// TIA Portal project "TestEssProtoFreia" (V13) (continued)

         AN    "ASCOenManuel";
         =     "PLC_to_Epics".CV550.sAuto;
END_REGION

REGION Network 13: spare - VB chan 7
   RUNG wire#powerrail
      Contact( "voie 7 chaufferette BV" )
      Coil( "PLC_to_Epics"."spare-VB-7".sHtrOn )
   END_RUNG
   // the same network as SCL:
   "PLC_to_Epics"."spare-VB-7".sHtrOn := "voie 7 chaufferette BV";
END_REGION

REGION Network 14: spare - VB chan 8
   RUNG wire#powerrail
      Contact( "voie 8 chaufferette BV" )
      Coil( "PLC_to_Epics"."spare-VB-8".sHtrOn )
   END_RUNG
   // the same network as SCL:
   "PLC_to_Epics"."spare-VB-8".sHtrOn := "voie 8 chaufferette BV";
END_REGION

REGION Network 15: spare VB chan 9
   RUNG wire#powerrail
      Contact( "voie 9 chaufferette BV" )
      Coil( "PLC_to_Epics"."spare-VB-9".sHtrOn )
   END_RUNG
   // the same network as SCL:
   "PLC_to_Epics"."spare-VB-9".sHtrOn := "voie 9 chaufferette BV";
END_REGION

REGION Network 16: spare - VB chan 10
   RUNG wire#powerrail
      Contact( "voie 10  chaufferette BV" )
      Coil( "PLC_to_Epics"."spare-VB-10".sHtrOn )
   END_RUNG
   // the same network as SCL:
   "PLC_to_Epics"."spare-VB-10".sHtrOn := "voie 10  chaufferette BV";
END_REGION

REGION Network 17: spare - VB chan 11
   RUNG wire#powerrail
      Contact( "voie 11 chaufferette BV" )
      Coil( "PLC_to_Epics"."spare-VB-11".sHtrOn )
   END_RUNG
   // the same network as SCL:
   "PLC_to_Epics"."spare-VB-11".sHtrOn := "voie 11 chaufferette BV";
END_REGION

REGION Network 18: EH901-902 CM chan 1
   RUNG wire#powerrail
      Contact( "voie 1 chaufferette CM" )
      Coil( "PLC_to_Epics"."EH901-902".sHtrOn )
   END_RUNG
   // the same network as SCL:
   "PLC_to_Epics"."EH901-902".sHtrOn := "voie 1 chaufferette CM";
END_REGION

REGION Network 19: EH913-914 CM channel 4
   RUNG wire#powerrail
      Contact( "voie 4 chaufferette CM" )
      Coil( "PLC_to_Epics"."EH913-914".sHtrOn )
   END_RUNG
   // the same network as SCL:
   "PLC_to_Epics"."EH913-914".sHtrOn := "voie 4 chaufferette CM";
END_REGION

REGION Network 20: EH933-934 - CM chan 5
   RUNG wire#powerrail
      Contact( "voie 5 chaufferette CM" )
      Coil( "PLC_to_Epics"."EH933-934".sHtrOn )
   END_RUNG
   // the same network as SCL:
   "PLC_to_Epics"."EH933-934".sHtrOn := "voie 5 chaufferette CM";
END_REGION

REGION Network 21: EH921 - CM chan 6
   RUNG wire#powerrail
      Contact( "voie 6 chaufferette CM" )
      Coil( "PLC_to_Epics".EH921.sHtrOn )
   END_RUNG
   // the same network as SCL:
   "PLC_to_Epics".EH921.sHtrOn := "voie 6 chaufferette CM";
END_REGION

REGION Network 22: EH931-932 - CM chan 7
   RUNG wire#powerrail
      Contact( "voie 7 chaufferette CM" )
      Coil( "PLC_to_Epics"."EH931-932".sHtrOn )
   END_RUNG
   // the same network as SCL:
   "PLC_to_Epics"."EH931-932".sHtrOn := "voie 7 chaufferette CM";
END_REGION

REGION Network 23: EH915-916 - CM chan 8
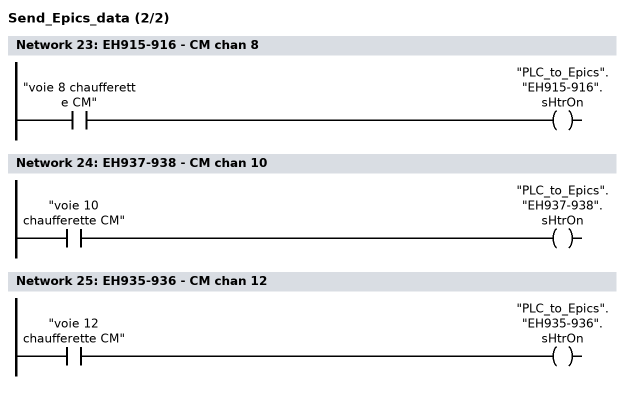
   RUNG wire#powerrail
      Contact( "voie 8 chaufferette CM" )
      Coil( "PLC_to_Epics"."EH915-916".sHtrOn )
   END_RUNG
   // the same network as SCL:
   "PLC_to_Epics"."EH915-916".sHtrOn := "voie 8 chaufferette CM";
END_REGION

REGION Network 24: EH937-938 - CM chan 10
   RUNG wire#powerrail
      Contact( "voie 10 chaufferette CM" )
      Coil( "PLC_to_Epics"."EH937-938".sHtrOn )
   END_RUNG
   // the same network as SCL:
   "PLC_to_Epics"."EH937-938".sHtrOn := "voie 10 chaufferette CM";
END_REGION

REGION Network 25: EH935-936 - CM chan 12
   RUNG wire#powerrail
      Contact( "voie 12 chaufferette CM" )
      Coil( "PLC_to_Epics"."EH935-936".sHtrOn )
   END_RUNG
   // the same network as SCL:
   "PLC_to_Epics"."EH935-936".sHtrOn := "voie 12 chaufferette CM";
END_REGION

REGION Network 26 (STL): Status bits
         A     "Graph/manuelle";
         =     "PLC_to_Epics".sManual;
         A     "ErreurSupervision";
         =     "PLC_to_Epics".sGrafcetERR;
         A     "Etat initial";
         =     "PLC_to_Epics".sGS1;
         A     "EtatCdtCryo";
         =     "PLC_to_Epics".sGS2;
         A     "EtatAttMef";
         =     "PLC_to_Epics".sGS3;
         A     "EtatMEFazote";
         =     "PLC_to_Epics".sGS4;
         A     "EtatMEFhelium";
         =     "PLC_to_Epics".sGS5;
         A     "EtatMode4k";
         =     "PLC_to_Epics".sGS6;
         A     "EtatModeStandBy";
         =     "PLC_to_Epics".sGS7;
         A     "EtatMode2K";
         =     "PLC_to_Epics".sGS8;
         A     "Etatrechauffage";
         =     "PLC_to_Epics".sGS10;
         A     "conditionTempMEFheliumOK";
         =     "PLC_to_Epics".sTransTempOK;
         A     "TransMode4K";
         =     "PLC_to_Epics".sTransMode4K;
         A     "EPICS_COMM_OK";
         =     "PLC_to_Epics".EpicsCommOK;
         A     "HNOSS_COMM_OK";
         =     "PLC_to_Epics".HNOSSCommOK;
END_REGION

REGION Network 27 (STL): Real parameters read-back (LHe level PID settings)
         L     "TriggerPIDcv01";
         T     "PLC_to_Epics".TrigPID_CV01.sSetV;
         L     "TriggerPIDcv02";
         T     "PLC_to_Epics".TrigPID_CV02.sSetV;
         L     "TriggerPIDcv03";
         T     "PLC_to_Epics".TrigPID_CV03.sSetV;
         L     "LT01LevelSP2k";
         T     "PLC_to_Epics".PID_LT01_CV01_SP.sSetV;
         L     "LT01LevelSP";
         T     "PLC_to_Epics".PID_LT01_CV02_SP.sSetV;
         L     "LT03LevelSP";
         T     "PLC_to_Epics".PID_LT03_CV03_SP.sSetV;
END_REGION

REGION Network 28 (STL): Real parameters read-back (CV550l PID settings)
         L     "RéguleASCO02_SP";
         T     "PLC_to_Epics".PID_PT01_CV550_SP.sSetV;
END_REGION
END_FUNCTION

FUNCTION "Cmds_from_Epics" : Void   // FC33, STL
TITLE = Process data from Epics
{ S7_Optimized_Access := 'FALSE' }
VERSION : 0.1
BEGIN

REGION Network 1: Switch to remote mode (control from Epics)
         A     "Epics_to_PLC".cmdRemoteMode;
         R     "LocalMode";
         R     "Epics_to_PLC".cmdRemoteMode;
END_REGION

REGION Network 2: If Local mode - return
         A     "LocalMode";
         SAVE;
         BEC;
END_REGION

REGION Network 3: Switch to local mode (control from Epics)
         A     "Epics_to_PLC".cmdLocalMode;
         S     "LocalMode";
         R     "Epics_to_PLC".cmdLocalMode;
END_REGION

REGION Network 4: If Local mode - return
         A     "LocalMode";
         SAVE;
         BEC;
END_REGION

REGION Network 5: Test data (copy block of data)
   //      OPN   "Epics_to_PLC"
   //      OPNDI "PLC_to_Epics"
   //      LAR1  P#12.0
   //      LAR2  P#12.0
   //      L     14
   //lp1:  T     #cnt
   //      L DBD [ AR1 , P#0.0 ]
   //      T DID [ AR2 , P#0.0 ]
   //      +AR1  P#4.0
   //      +AR2  P#4.0
   //      L     #cnt
   //      LOOP  lp1
END_REGION

REGION Network 6: CV01 Man/Auto
         A     "Epics_to_PLC".CV01.cmdAuto;
         R     "CV01_ManAuto";
         A     "Epics_to_PLC".CV01.cmdMan;
         S     "CV01_ManAuto";
END_REGION

REGION Network 7: CV01 - set Value
         A     "CV01_ManAuto";
         A     "Epics_to_PLC".CV01.cmdSet;
         JNB   Label_0;
         L     "Epics_to_PLC".CV01.cSetv;
         T     "CV01_HMI_VAL";
         SET;
         SAVE;
         CLR;
   Label_0:A     BR;
         R     "Epics_to_PLC".CV01.cmdSet;
END_REGION

REGION Network 8: CV02 Man/Auto
         A     "Epics_to_PLC".CV02.cmdAuto;
         R     "CV02_ManAuto";
         A     "Epics_to_PLC".CV02.cmdMan;
         S     "CV02_ManAuto";
END_REGION

REGION Network 9: CV02 - set Value
         A     "CV02_ManAuto";
         A     "Epics_to_PLC".CV02.cmdSet;
         JNB   Label_1;
         L     "Epics_to_PLC".CV02.cSetv;
         T     "CV02_HMI_VAL";
         SET;
         SAVE;
         CLR;
   Label_1:A     BR;
         R     "Epics_to_PLC".CV02.cmdSet;
END_REGION

REGION Network 10: CV03 Man/Auto
         A     "Epics_to_PLC".CV03.cmdAuto;
         R     "CV03_ManAuto";
         A     "Epics_to_PLC".CV03.cmdMan;
         S     "CV03_ManAuto";
END_REGION

REGION Network 11: CV03 - set Value
         A     "CV03_ManAuto";
         A     "Epics_to_PLC".CV03.cmdSet;
         JNB   Label_2;
         L     "Epics_to_PLC".CV03.cSetv;
         T     "CV03_HMI_VAL";
         SET;
         SAVE;
         CLR;
   Label_2:A     BR;
         R     "Epics_to_PLC".CV03.cmdSet;
END_REGION

REGION Network 12: CV04 Man/Auto
         A     "Epics_to_PLC".CV04.cmdAuto;
         R     "CV04_ManAuto";
         A     "Epics_to_PLC".CV04.cmdMan;
         S     "CV04_ManAuto";
END_REGION

REGION Network 13: CV04 - set Value
         A     "CV04_ManAuto";
         A     "Epics_to_PLC".CV04.cmdSet;
         JNB   Label_3;
         L     "Epics_to_PLC".CV04.cSetv;
         T     "CV04_HMI_VAL";
         SET;
         SAVE;
         CLR;
   Label_3:A     BR;
         R     "Epics_to_PLC".CV04.cmdSet;
END_REGION

REGION Network 14: CV05 Man/Auto
END_REGION

REGION Network 15: CV05 - set Value NOTE: NO LOCAL FALG !!!!!!!!!!!!!!!!!!!
         A     "Epics_to_PLC".CV05.cmdSet;
         JNB   Label_4;
         L     "Epics_to_PLC".CV05.cSetv;
         T     "CV05_HMI_VAL";
         SET;
         SAVE;
         CLR;
   Label_4:A     BR;
         R     "Epics_to_PLC".CV05.cmdSet;
END_REGION

REGION Network 16: CV07 Man/Auto
         A     "Epics_to_PLC".CV07.cmdAuto;
         R     "CV07_ManAuto";
         A     "Epics_to_PLC".CV07.cmdMan;
         S     "CV07_ManAuto";
END_REGION

REGION Network 17: CV07 - set Value
         A     "CV07_ManAuto";
         A     "Epics_to_PLC".CV07.cmdSet;
         JNB   Label_5;
         L     "Epics_to_PLC".CV07.cSetv;
         T     "CV07_HMI_VAL";
         SET;
         SAVE;
         CLR;
   Label_5:A     BR;
         R     "Epics_to_PLC".CV07.cmdSet;
END_REGION

REGION Network 18: CV60 Man/Auto
         A     "Epics_to_PLC".CV60.cmdAuto;
         R     "CV60_ManAuto";
         A     "Epics_to_PLC".CV60.cmdMan;
         S     "CV60_ManAuto";
END_REGION

REGION Network 19: CV60 - set Value
         A     "CV60_ManAuto";
         A     "Epics_to_PLC".CV60.cmdSet;
         JNB   Label_6;
         L     "Epics_to_PLC".CV60.cSetv;
         T     "CV60_HMI_VAL";
         SET;
         SAVE;
         CLR;
   Label_6:A     BR;
         R     "Epics_to_PLC".CV60.cmdSet;
END_REGION

REGION Network 20: CV61 Man/Auto
         A     "Epics_to_PLC".CV61.cmdAuto;
         R     "CV61_ManAuto";
         A     "Epics_to_PLC".CV61.cmdMan;
         S     "CV61_ManAuto";
END_REGION

REGION Network 21: CV61 - set Value
         A     "CV61_ManAuto";
         A     "Epics_to_PLC".CV61.cmdSet;
         JNB   Label_7;
         L     "Epics_to_PLC".CV61.cSetv;
         T     "CV61_HMI_VAL";
         SET;
         SAVE;
         CLR;
   Label_7:A     BR;
         R     "Epics_to_PLC".CV61.cmdSet;
END_REGION

REGION Network 22: CV62 Man/Auto
END_REGION

REGION Network 23: CV62 - set Value
         A     "Epics_to_PLC".CV62.cmdSet;
         JNB   Label_8;
         L     "Epics_to_PLC".CV62.cSetv;
         T     "CV62_HMI_VAL";
         SET;
         SAVE;
         CLR;
   Label_8:A     BR;
         R     "Epics_to_PLC".CV62.cmdSet;
END_REGION

REGION Network 24: CV550 Man/Auto
         A     "Epics_to_PLC".CV550.cmdAuto;
         R     "ASCOenManuel";
         A     "Epics_to_PLC".CV550.cmdMan;
         S     "ASCOenManuel";
END_REGION

REGION Network 25: CV550 - set Value
         A     "ASCOenManuel";
         A     "Epics_to_PLC".CV550.cmdSet;
         JNB   Label_9;
         L     "Epics_to_PLC".CV550.cSetv;
         T     "Asco02ManValeur";
         SET;
         SAVE;
         CLR;
   Label_9:A     BR;
         R     "Epics_to_PLC".CV550.cmdSet;
END_REGION

REGION Network 26: spare- VB chan 7
         A     "Epics_to_PLC"."spare-VB-7".cmdSet;
         S     "voie 7 chaufferette BV";
         A     "Epics_to_PLC"."spare-VB-7".cmdRst;
         R     "voie 7 chaufferette BV";
END_REGION

REGION Network 27: spare- VB chan 8
         A     "Epics_to_PLC"."spare-VB-8".cmdSet;
         S     "voie 8 chaufferette BV";
         A     "Epics_to_PLC"."spare-VB-8".cmdRst;
         R     "voie 8 chaufferette BV";
END_REGION

REGION Network 28: spare- VB chan 9
         A     "Epics_to_PLC"."spare-VB-9".cmdSet;
         S     "voie 9 chaufferette BV";
         A     "Epics_to_PLC"."spare-VB-9".cmdRst;
         R     "voie 9 chaufferette BV";
END_REGION

REGION Network 29: spare- VB chan 10
         A     "Epics_to_PLC"."spare-VB-10".cmdSet;
         S     "voie 10  chaufferette BV";
         A     "Epics_to_PLC"."spare-VB-10".cmdRst;
         R     "voie 10  chaufferette BV";
END_REGION

REGION Network 30: spare - VB chan 11
         A     "Epics_to_PLC"."spare-VB-11".cmdSet;
         S     "voie 11 chaufferette BV";
         A     "Epics_to_PLC"."spare-VB-11".cmdRst;
         R     "voie 11 chaufferette BV";
END_REGION

REGION Network 31: EH901-902 CM chan 1
         A     "Epics_to_PLC"."EH901-902".cmdSet;
         S     "voie 1 chaufferette CM";
         A     "Epics_to_PLC"."EH901-902".cmdRst;
         R     "voie 1 chaufferette CM";
END_REGION

REGION Network 32: EH913-914 CM chan 4
         A     "Epics_to_PLC"."EH913-914".cmdSet;
         S     "voie 4 chaufferette CM";
         A     "Epics_to_PLC"."EH913-914".cmdRst;
         R     "voie 4 chaufferette CM";
END_REGION

REGION Network 33: EH933-934 - CM chan 5
         A     "Epics_to_PLC"."EH933-934".cmdSet;
         S     "voie 5 chaufferette CM";
         A     "Epics_to_PLC"."EH933-934".cmdRst;
         R     "voie 5 chaufferette CM";
END_REGION

REGION Network 34: EH921 - CM chan 6
         A     "Epics_to_PLC".EH921.cmdSet;
         S     "voie 6 chaufferette CM";
         A     "Epics_to_PLC".EH921.cmdRst;
         R     "voie 6 chaufferette CM";
END_REGION

REGION Network 35: EH931-932 - CM chan 7
         A     "Epics_to_PLC"."EH931-932".cmdSet;
         S     "voie 7 chaufferette CM";
         A     "Epics_to_PLC"."EH931-932".cmdRst;
         R     "voie 7 chaufferette CM";
END_REGION

REGION Network 36: EH915-916 - CM chan 8
         A     "Epics_to_PLC"."EH915-916".cmdSet;
         S     "voie 8 chaufferette CM";
         A     "Epics_to_PLC"."EH915-916".cmdRst;
         R     "voie 8 chaufferette CM";
END_REGION

REGION Network 37: EH937-938 - CM chan 10
         A     "Epics_to_PLC"."EH937-938".cmdSet;
         S     "voie 10 chaufferette CM";
         A     "Epics_to_PLC"."EH937-938".cmdRst;
         R     "voie 10 chaufferette CM";
END_REGION

REGION Network 38: EH935-936 - CM chan 12
         A     "Epics_to_PLC"."EH935-936".cmdSet;
         S     "voie 12 chaufferette CM";
         A     "Epics_to_PLC"."EH935-936".cmdRst;
         R     "voie 12 chaufferette CM";
END_REGION

REGION Network 39: Bit commands
         A     "Epics_to_PLC".cmdAutoMode;
         R     "Graph/manuelle";
         A     "Epics_to_PLC".cmdManMode;
         S     "Graph/manuelle";
         A     "Epics_to_PLC".cmdGrafcetInit;
         =     "MettreEtatInitial";
         A     "Epics_to_PLC".cmdGrafcetErrRst;
         =     "AcquitterErreurGraph";
         A     "Epics_to_PLC".cmdStartConditioning;
         =     "CmdVanneEtatCdt";
         A     "Epics_to_PLC".cmdCondOK;
         =     "CdtInfraOk";
         A     "Epics_to_PLC".cmdCondERR;
         =     "CdtInfraErreur";
         A     "Epics_to_PLC".cmdStartLN2cooling;
         =     "DmdMefAzote";
         A     "Epics_to_PLC".cmdStartLHecooling;
         =     "DmdMefHelium";
         A     "Epics_to_PLC".cmdStart2Kmode;
         =     "DmdMode2K";
         A     "Epics_to_PLC".cmdStop2Kmode;
         =     "DmdArretMode2k";
         A     "Epics_to_PLC".cmdStartSTBYmode;
         =     "DmdModeStandby";
         A     "Epics_to_PLC".cmdStopSTBYmode;
         =     "DmdArretModeStandby";
         A     "Epics_to_PLC".cmdStartHeating;
         =     "StartHeating";
         A     "Epics_to_PLC".cmdStopHeating;
         =     "StopHeating";
END_REGION

REGION Network 40: Real parameters (LHe level PIDs settings)
         A     "Epics_to_PLC".TrigPID_CV01.cmdSet;
         JNB   Label_10;
         L     "Epics_to_PLC".TrigPID_CV01.cSetV;
         T     "TriggerPIDcv01";
         SET;
         SAVE;
         CLR;
   Label_10:A     BR;
         R     "Epics_to_PLC".TrigPID_CV01.cmdSet;
END_REGION

REGION Network 41: Real parameters (LHe level PIDs settings)
         A     "Epics_to_PLC".TrigPID_CV02.cmdSet;
         JNB   Label_11;
         L     "Epics_to_PLC".TrigPID_CV02.cSetV;
         T     "TriggerPIDcv02";
         SET;
         SAVE;
         CLR;
   Label_11:A     BR;
         R     "Epics_to_PLC".TrigPID_CV02.cmdSet;
END_REGION

REGION Network 42: Real parameters (LHe level PIDs settings)
         A     "Epics_to_PLC".TrigPID_CV03.cmdSet;
         JNB   Label_12;
         L     "Epics_to_PLC".TrigPID_CV03.cSetV;
         T     "TriggerPIDcv03";
         SET;
         SAVE;
         CLR;
   Label_12:A     BR;
         R     "Epics_to_PLC".TrigPID_CV03.cmdSet;
END_REGION

REGION Network 43: Real parameters (LHe level PIDs settings)
         A     "Epics_to_PLC".PID_LT01_CV01_SP.cmdSet;
         JNB   Label_13;
         L     "Epics_to_PLC".PID_LT01_CV01_SP.cSetV;
         T     "LT01LevelSP2k";
         SET;
         SAVE;
         CLR;
   Label_13:A     BR;
         R     "Epics_to_PLC".PID_LT01_CV01_SP.cmdSet;
END_REGION

REGION Network 44: Real parameters (LHe level PIDs settings)
         A     "Epics_to_PLC".PID_LT03_CV03_SP.cmdSet;
         JNB   Label_14;
         L     "Epics_to_PLC".PID_LT03_CV03_SP.cSetV;
         T     "LT03LevelSP";
         SET;
         SAVE;
         CLR;
   Label_14:A     BR;
         R     "Epics_to_PLC".PID_LT03_CV03_SP.cmdSet;
END_REGION

REGION Network 45: Real parameters (LHe level PIDs settings)
         A     "Epics_to_PLC".PID_LT01_CV02_SP.cmdSet;
         JNB   Label_16;
         L     "Epics_to_PLC".PID_LT01_CV02_SP.cSetV;
         T     "LT01LevelSP";
         SET;
         SAVE;
         CLR;
   Label_16:A     BR;

         R     "Epics_to_PLC".PID_LT01_CV02_SP.cmdSet;
END_REGION

REGION Network 46: Real parameters (PT01 PIDs settings)
         A     "Epics_to_PLC".PID_PT01_CV550_SP.cmdSet;
         JNB   Label_15;
         L     "Epics_to_PLC".PID_PT01_CV550_SP.cSetV;
         T     "RéguleASCO02_SP";
         SET;
         SAVE;
         CLR;
   Label_15:A     BR;
         R     "Epics_to_PLC".PID_PT01_CV550_SP.cmdSet;
END_REGION

REGION Network 47: Temperatures fromKeithley
         L     "Epics_to_PLC".TTxx;
         T     "ReceivePT100"."TTxx_(K)";
         L     "Epics_to_PLC".TTyy;
         T     "ReceivePT100"."TTyy_(K)";
END_REGION
END_FUNCTION

FUNCTION "Data_from_IOC" : Void   // FC34, LAD
TITLE = Get data from the IOC andcheck if the connection is alive
{ S7_Optimized_Access := 'FALSE' }
VERSION : 0.1
BEGIN

REGION Network 1: Check the Data from the IOC
END_REGION
END_FUNCTION

FUNCTION "grafcet" : Void   // FC99, LAD
{ S7_Optimized_Access := 'FALSE' }
VERSION : 0.1
   VAR_TEMP   // added for the SCL form of the ladder/FBD networks
      _w1 : Bool;
      _w2 : Bool;
      _w3 : Bool;
      _w4 : Bool;
      _w5 : Bool;
      _w6 : Bool;
      _w7 : Bool;
      _w8 : Bool;
   END_VAR
BEGIN

REGION Network 1: config vannes init mode
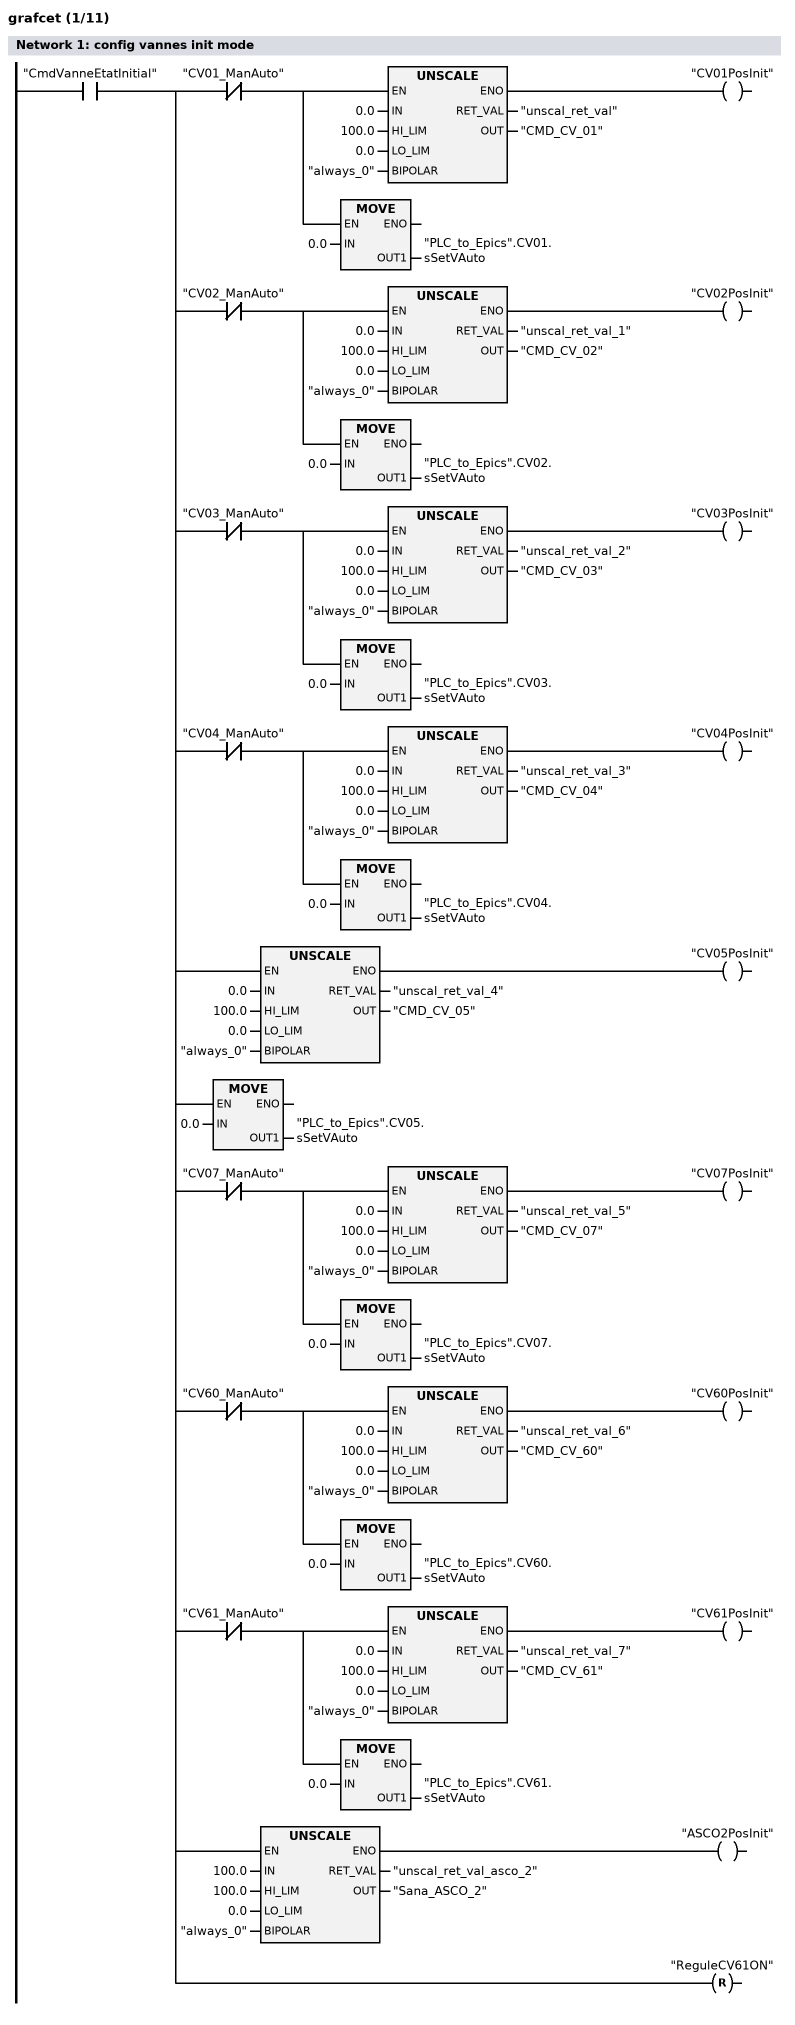
   // ENO of a box is taken as its EN; it also drops when the box reports an error
   #_w1 := "CmdVanneEtatInitial" AND NOT "CV01_ManAuto";
   #_w2 := "CmdVanneEtatInitial";
   IF #_w1 THEN
       "unscal_ret_val" := UNSCALE(IN := 0.0,
                               HI_LIM := 100.0,
                               LO_LIM := 0.0,
                               BIPOLAR := "always_0",
                               OUT => "CMD_CV_01");
   END_IF;
   "CV01PosInit" := #_w1;
   IF #_w1 THEN "PLC_to_Epics".CV01.sSetVAuto := 0.0; END_IF;
   #_w3 := #_w2 AND NOT "CV02_ManAuto";
   IF #_w3 THEN
       "unscal_ret_val_1" := UNSCALE(IN := 0.0,
                               HI_LIM := 100.0,
                               LO_LIM := 0.0,
                               BIPOLAR := "always_0",
                               OUT => "CMD_CV_02");
   END_IF;
   "CV02PosInit" := #_w3;
   IF #_w3 THEN "PLC_to_Epics".CV02.sSetVAuto := 0.0; END_IF;
   #_w4 := #_w2 AND NOT "CV03_ManAuto";
   IF #_w4 THEN
       "unscal_ret_val_2" := UNSCALE(IN := 0.0,
                               HI_LIM := 100.0,
                               LO_LIM := 0.0,
                               BIPOLAR := "always_0",
                               OUT => "CMD_CV_03");
   END_IF;
   "CV03PosInit" := #_w4;
   IF #_w4 THEN "PLC_to_Epics".CV03.sSetVAuto := 0.0; END_IF;
   #_w5 := #_w2 AND NOT "CV04_ManAuto";
   IF #_w5 THEN
       "unscal_ret_val_3" := UNSCALE(IN := 0.0,
                               HI_LIM := 100.0,
                               LO_LIM := 0.0,
                               BIPOLAR := "always_0",
                               OUT => "CMD_CV_04");
   END_IF;
   "CV04PosInit" := #_w5;
   IF #_w5 THEN "PLC_to_Epics".CV04.sSetVAuto := 0.0; END_IF;
   IF #_w2 THEN
       "unscal_ret_val_4" := UNSCALE(IN := 0.0,
                               HI_LIM := 100.0,
                               LO_LIM := 0.0,
                               BIPOLAR := "always_0",
                               OUT => "CMD_CV_05");
   END_IF;
   "CV05PosInit" := #_w2;
   IF #_w2 THEN "PLC_to_Epics".CV05.sSetVAuto := 0.0; END_IF;
   #_w6 := #_w2 AND NOT "CV07_ManAuto";
   IF #_w6 THEN
       "unscal_ret_val_5" := UNSCALE(IN := 0.0,
                               HI_LIM := 100.0,
                               LO_LIM := 0.0,
                               BIPOLAR := "always_0",
                               OUT => "CMD_CV_07");
   END_IF;
   "CV07PosInit" := #_w6;
   IF #_w6 THEN "PLC_to_Epics".CV07.sSetVAuto := 0.0; END_IF;
   #_w7 := #_w2 AND NOT "CV60_ManAuto";
   IF #_w7 THEN
       "unscal_ret_val_6" := UNSCALE(IN := 0.0,
                               HI_LIM := 100.0,
                               LO_LIM := 0.0,
                               BIPOLAR := "always_0",
                               OUT => "CMD_CV_60");
   END_IF;
   "CV60PosInit" := #_w7;
   IF #_w7 THEN "PLC_to_Epics".CV60.sSetVAuto := 0.0; END_IF;
   #_w8 := #_w2 AND NOT "CV61_ManAuto";
   IF #_w8 THEN
       "unscal_ret_val_7" := UNSCALE(IN := 0.0,
                               HI_LIM := 100.0,
                               LO_LIM := 0.0,
                               BIPOLAR := "always_0",
                               OUT => "CMD_CV_61");
   END_IF;
   "CV61PosInit" := #_w8;
   IF #_w8 THEN "PLC_to_Epics".CV61.sSetVAuto := 0.0; END_IF;
   IF #_w2 THEN
       "unscal_ret_val_asco_2" := UNSCALE(IN := 100.0,
                               HI_LIM := 100.0,
                               LO_LIM := 0.0,
                               BIPOLAR := "always_0",
                               OUT => "Sana_ASCO_2");
   END_IF;
   "ASCO2PosInit" := #_w2;
   IF #_w2 THEN "ReguleCV61ON" := FALSE; END_IF;
END_REGION

REGION Network 2: Vanne En Position Initial
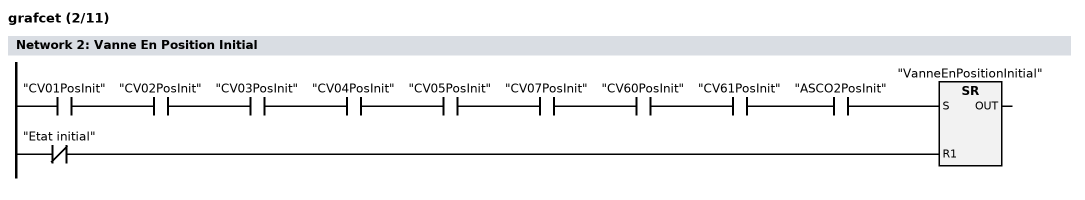
   RUNG wire#powerrail
      Contact( "CV01PosInit" )
      Contact( "CV02PosInit" )
      Contact( "CV03PosInit" )
      Contact( "CV04PosInit" )
      Contact( "CV05PosInit" )
      Contact( "CV07PosInit" )
      Contact( "CV60PosInit" )
      Contact( "CV61PosInit" )
      Contact( "ASCO2PosInit" )
      S_SR(operand := "VanneEnPositionInitial", r1 := wire#w1)
   END_RUNG
   RUNG wire#powerrail
      I_Contact( "Etat initial" )
   END_RUNG wire#w1
   // the same network as SCL:
   IF "CV01PosInit" AND "CV02PosInit" AND "CV03PosInit" AND "CV04PosInit" AND "CV05PosInit" AND "CV07PosInit" AND "CV60PosInit" AND "CV61PosInit" AND "ASCO2PosInit" THEN
       "VanneEnPositionInitial" := TRUE;   // SR flip-flop
   END_IF;
   IF NOT "Etat initial" THEN "VanneEnPositionInitial" := FALSE; END_IF;
END_REGION

REGION Network 3: config vanne etat conditionnement
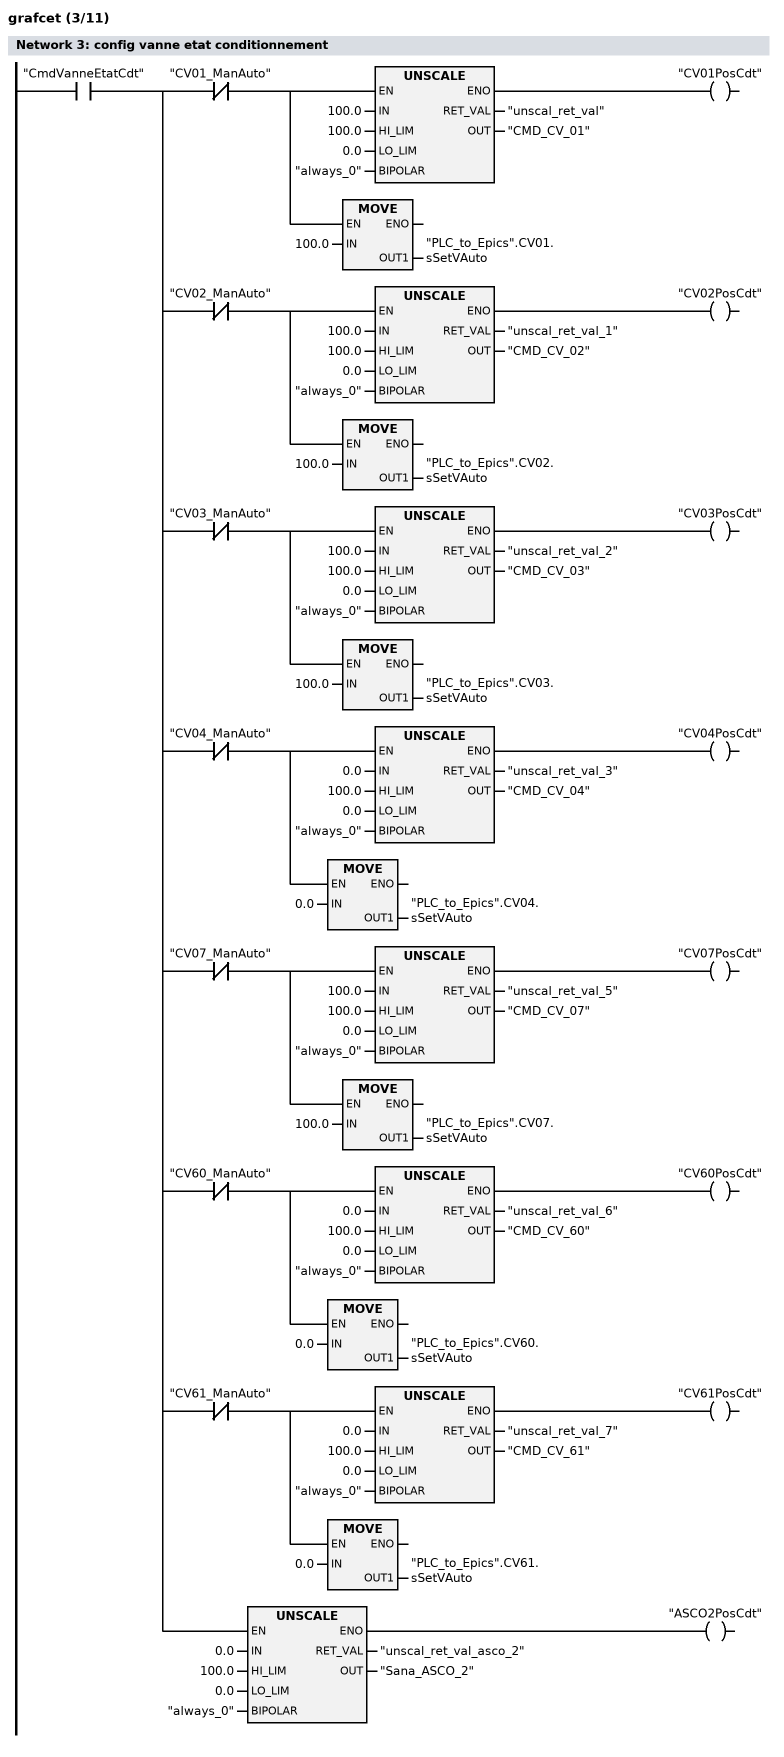
   // ENO of a box is taken as its EN; it also drops when the box reports an error
   #_w1 := "CmdVanneEtatCdt" AND NOT "CV01_ManAuto";
   #_w2 := "CmdVanneEtatCdt";
   IF #_w1 THEN
       "unscal_ret_val" := UNSCALE(IN := 100.0,
                               HI_LIM := 100.0,
                               LO_LIM := 0.0,
                               BIPOLAR := "always_0",
                               OUT => "CMD_CV_01");
   END_IF;
   "CV01PosCdt" := #_w1;
   IF #_w1 THEN "PLC_to_Epics".CV01.sSetVAuto := 100.0; END_IF;
   #_w3 := #_w2 AND NOT "CV02_ManAuto";
   IF #_w3 THEN
       "unscal_ret_val_1" := UNSCALE(IN := 100.0,
                               HI_LIM := 100.0,
                               LO_LIM := 0.0,
                               BIPOLAR := "always_0",
                               OUT => "CMD_CV_02");
   END_IF;
   "CV02PosCdt" := #_w3;
   IF #_w3 THEN "PLC_to_Epics".CV02.sSetVAuto := 100.0; END_IF;
   #_w4 := #_w2 AND NOT "CV03_ManAuto";
   IF #_w4 THEN
       "unscal_ret_val_2" := UNSCALE(IN := 100.0,
                               HI_LIM := 100.0,
                               LO_LIM := 0.0,
                               BIPOLAR := "always_0",
                               OUT => "CMD_CV_03");
   END_IF;
   "CV03PosCdt" := #_w4;
   IF #_w4 THEN "PLC_to_Epics".CV03.sSetVAuto := 100.0; END_IF;
   #_w5 := #_w2 AND NOT "CV04_ManAuto";
   IF #_w5 THEN
       "unscal_ret_val_3" := UNSCALE(IN := 0.0,
                               HI_LIM := 100.0,
                               LO_LIM := 0.0,
                               BIPOLAR := "always_0",
                               OUT => "CMD_CV_04");
   END_IF;
   "CV04PosCdt" := #_w5;
   IF #_w5 THEN "PLC_to_Epics".CV04.sSetVAuto := 0.0; END_IF;
   #_w6 := #_w2 AND NOT "CV07_ManAuto";
   IF #_w6 THEN
       "unscal_ret_val_5" := UNSCALE(IN := 100.0,
                               HI_LIM := 100.0,
                               LO_LIM := 0.0,
                               BIPOLAR := "always_0",
                               OUT => "CMD_CV_07");
   END_IF;
   "CV07PosCdt" := #_w6;
   IF #_w6 THEN "PLC_to_Epics".CV07.sSetVAuto := 100.0; END_IF;
   #_w7 := #_w2 AND NOT "CV60_ManAuto";
   IF #_w7 THEN
       "unscal_ret_val_6" := UNSCALE(IN := 0.0,
                               HI_LIM := 100.0,
                               LO_LIM := 0.0,
                               BIPOLAR := "always_0",
                               OUT => "CMD_CV_60");
   END_IF;
   "CV60PosCdt" := #_w7;
   IF #_w7 THEN "PLC_to_Epics".CV60.sSetVAuto := 0.0; END_IF;
   #_w8 := #_w2 AND NOT "CV61_ManAuto";
   IF #_w8 THEN
       "unscal_ret_val_7" := UNSCALE(IN := 0.0,
                               HI_LIM := 100.0,
                               LO_LIM := 0.0,
                               BIPOLAR := "always_0",
                               OUT => "CMD_CV_61");
   END_IF;
   "CV61PosCdt" := #_w8;
   IF #_w8 THEN "PLC_to_Epics".CV61.sSetVAuto := 0.0; END_IF;
   IF #_w2 THEN
       "unscal_ret_val_asco_2" := UNSCALE(IN := 0.0,
                               HI_LIM := 100.0,
                               LO_LIM := 0.0,
                               BIPOLAR := "always_0",
                               OUT => "Sana_ASCO_2");
   END_IF;
   "ASCO2PosCdt" := #_w2;
END_REGION

REGION Network 4: Vanne En Position Cdt
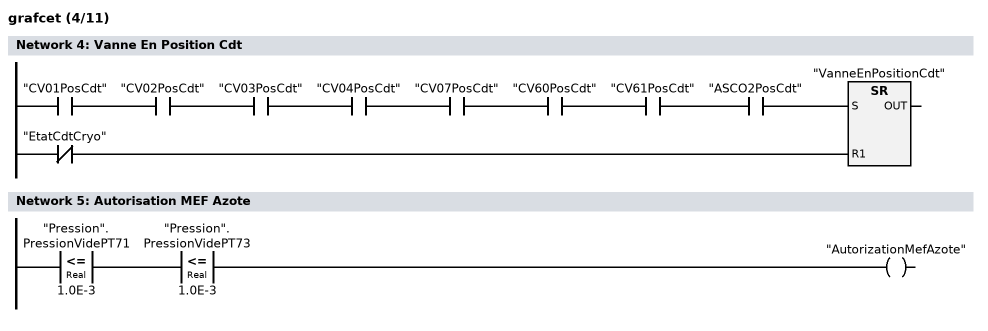
   RUNG wire#powerrail
      Contact( "CV01PosCdt" )
      Contact( "CV02PosCdt" )
      Contact( "CV03PosCdt" )
      Contact( "CV04PosCdt" )
      Contact( "CV07PosCdt" )
      Contact( "CV60PosCdt" )
      Contact( "CV61PosCdt" )
      Contact( "ASCO2PosCdt" )
      S_SR(operand := "VanneEnPositionCdt", r1 := wire#w1)
   END_RUNG
   RUNG wire#powerrail
      I_Contact( "EtatCdtCryo" )
   END_RUNG wire#w1
   // the same network as SCL:
   IF "CV01PosCdt" AND "CV02PosCdt" AND "CV03PosCdt" AND "CV04PosCdt" AND "CV07PosCdt" AND "CV60PosCdt" AND "CV61PosCdt" AND "ASCO2PosCdt" THEN
       "VanneEnPositionCdt" := TRUE;   // SR flip-flop
   END_IF;
   IF NOT "EtatCdtCryo" THEN "VanneEnPositionCdt" := FALSE; END_IF;
END_REGION

REGION Network 5: Autorisation MEF Azote
   RUNG wire#powerrail
      { S7_Templates := "SrcType := Real" } LE_Contact(in1 := "Pression".PressionVidePT71, in2 := 1.0E-3)
      { S7_Templates := "SrcType := Real" } LE_Contact(in1 := "Pression".PressionVidePT73, in2 := 1.0E-3)
      Coil( "AutorizationMefAzote" )
   END_RUNG
   // the same network as SCL:
   "AutorizationMefAzote" := ("Pression".PressionVidePT71 <= 1.0E-3) AND ("Pression".PressionVidePT73 <= 1.0E-3);
END_REGION

REGION Network 6: config vannes init mode & regule cv61 on
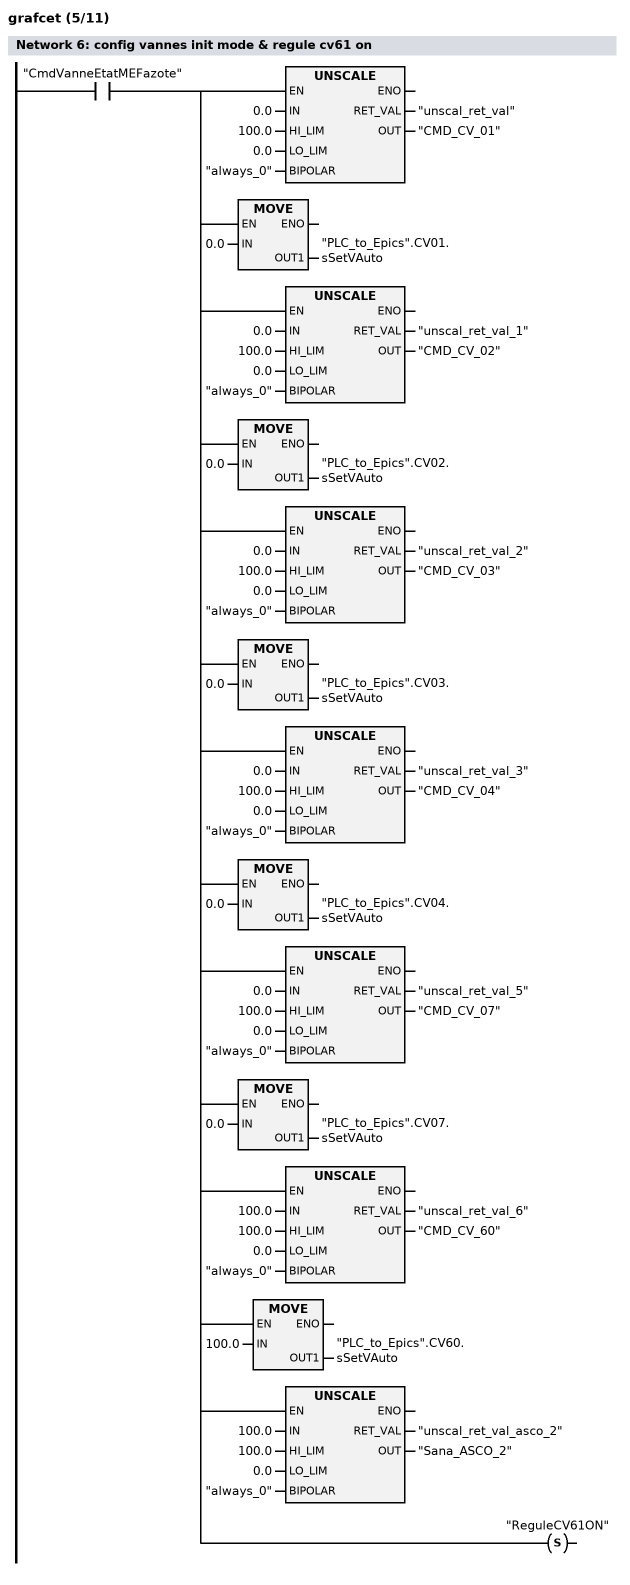
   #_w1 := "CmdVanneEtatMEFazote";
   IF #_w1 THEN
       "unscal_ret_val" := UNSCALE(IN := 0.0,
                               HI_LIM := 100.0,
                               LO_LIM := 0.0,
                               BIPOLAR := "always_0",
                               OUT => "CMD_CV_01");
       "PLC_to_Epics".CV01.sSetVAuto := 0.0;
       "unscal_ret_val_1" := UNSCALE(IN := 0.0,
                               HI_LIM := 100.0,
                               LO_LIM := 0.0,
                               BIPOLAR := "always_0",
                               OUT => "CMD_CV_02");
       "PLC_to_Epics".CV02.sSetVAuto := 0.0;
       "unscal_ret_val_2" := UNSCALE(IN := 0.0,
                               HI_LIM := 100.0,
                               LO_LIM := 0.0,
                               BIPOLAR := "always_0",
                               OUT => "CMD_CV_03");
       "PLC_to_Epics".CV03.sSetVAuto := 0.0;
       "unscal_ret_val_3" := UNSCALE(IN := 0.0,
                               HI_LIM := 100.0,
                               LO_LIM := 0.0,
                               BIPOLAR := "always_0",
                               OUT => "CMD_CV_04");
       "PLC_to_Epics".CV04.sSetVAuto := 0.0;
       "unscal_ret_val_5" := UNSCALE(IN := 0.0,
                               HI_LIM := 100.0,
                               LO_LIM := 0.0,
                               BIPOLAR := "always_0",
                               OUT => "CMD_CV_07");
       "PLC_to_Epics".CV07.sSetVAuto := 0.0;
       "unscal_ret_val_6" := UNSCALE(IN := 100.0,
                               HI_LIM := 100.0,
                               LO_LIM := 0.0,
                               BIPOLAR := "always_0",
                               OUT => "CMD_CV_60");
       "PLC_to_Epics".CV60.sSetVAuto := 100.0;
       "unscal_ret_val_asco_2" := UNSCALE(IN := 100.0,
                               HI_LIM := 100.0,
                               LO_LIM := 0.0,
                               BIPOLAR := "always_0",
                               OUT => "Sana_ASCO_2");
       "ReguleCV61ON" := TRUE;
   END_IF;
END_REGION

